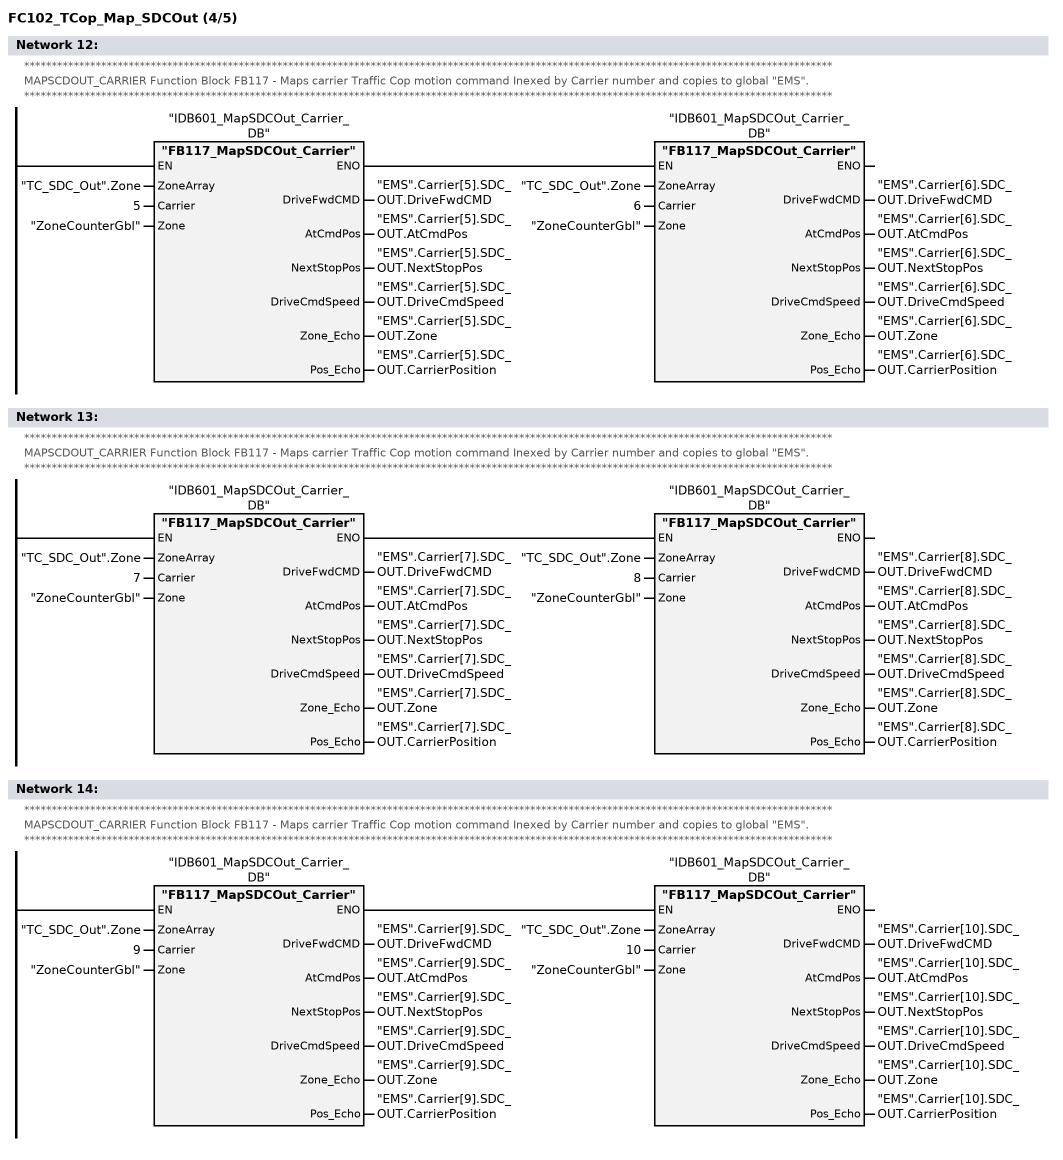
   RUNG wire#powerrail
      "IDB601_MapSDCOut_Carrier_DB"(ZoneArray := "TC_SDC_Out".Zone, Carrier := 5, Zone := "ZoneCounterGbl", DriveFwdCMD => "EMS".Carrier[5].SDC_OUT.DriveFwdCMD, AtCmdPos => "EMS".Carrier[5].SDC_OUT.AtCmdPos, NextStopPos => "EMS".Carrier[5].SDC_OUT.NextStopPos, DriveCmdSpeed => "EMS".Carrier[5].SDC_OUT.DriveCmdSpeed, Zone_Echo => "EMS".Carrier[5].SDC_OUT.Zone, Pos_Echo => "EMS".Carrier[5].SDC_OUT.CarrierPosition)
      "IDB601_MapSDCOut_Carrier_DB"(ZoneArray := "TC_SDC_Out".Zone, Carrier := 6, Zone := "ZoneCounterGbl", DriveFwdCMD => "EMS".Carrier[6].SDC_OUT.DriveFwdCMD, AtCmdPos => "EMS".Carrier[6].SDC_OUT.AtCmdPos, NextStopPos => "EMS".Carrier[6].SDC_OUT.NextStopPos, DriveCmdSpeed => "EMS".Carrier[6].SDC_OUT.DriveCmdSpeed, Zone_Echo => "EMS".Carrier[6].SDC_OUT.Zone, Pos_Echo => "EMS".Carrier[6].SDC_OUT.CarrierPosition)
   END_RUNG
   // the same network as SCL:
   "IDB601_MapSDCOut_Carrier_DB"(ZoneArray := "TC_SDC_Out".Zone,   // "FB117_MapSDCOut_Carrier"
                           Carrier := 5,
                           Zone := "ZoneCounterGbl",
                           DriveFwdCMD => "EMS".Carrier[5].SDC_OUT.DriveFwdCMD,
                           AtCmdPos => "EMS".Carrier[5].SDC_OUT.AtCmdPos,
                           NextStopPos => "EMS".Carrier[5].SDC_OUT.NextStopPos,
                           DriveCmdSpeed => "EMS".Carrier[5].SDC_OUT.DriveCmdSpeed,
                           Zone_Echo => "EMS".Carrier[5].SDC_OUT.Zone,
                           Pos_Echo => "EMS".Carrier[5].SDC_OUT.CarrierPosition,
                           ENO => #_w1);
   IF #_w1 THEN
       "IDB601_MapSDCOut_Carrier_DB"(ZoneArray := "TC_SDC_Out".Zone,   // "FB117_MapSDCOut_Carrier"
                               Carrier := 6,
                               Zone := "ZoneCounterGbl",
                               DriveFwdCMD => "EMS".Carrier[6].SDC_OUT.DriveFwdCMD,
                               AtCmdPos => "EMS".Carrier[6].SDC_OUT.AtCmdPos,
                               NextStopPos => "EMS".Carrier[6].SDC_OUT.NextStopPos,
                               DriveCmdSpeed => "EMS".Carrier[6].SDC_OUT.DriveCmdSpeed,
                               Zone_Echo => "EMS".Carrier[6].SDC_OUT.Zone,
                               Pos_Echo => "EMS".Carrier[6].SDC_OUT.CarrierPosition);
   END_IF;
END_REGION

REGION Network 13
   // ***************************************************************************************************************************************************
   // 
   // MAPSCDOUT_CARRIER Function Block FB117 - Maps carrier Traffic Cop motion command Inexed by Carrier number and copies to global "EMS". 
   // 
   // ***************************************************************************************************************************************************
   RUNG wire#powerrail
      "IDB601_MapSDCOut_Carrier_DB"(ZoneArray := "TC_SDC_Out".Zone, Carrier := 7, Zone := "ZoneCounterGbl", DriveFwdCMD => "EMS".Carrier[7].SDC_OUT.DriveFwdCMD, AtCmdPos => "EMS".Carrier[7].SDC_OUT.AtCmdPos, NextStopPos => "EMS".Carrier[7].SDC_OUT.NextStopPos, DriveCmdSpeed => "EMS".Carrier[7].SDC_OUT.DriveCmdSpeed, Zone_Echo => "EMS".Carrier[7].SDC_OUT.Zone, Pos_Echo => "EMS".Carrier[7].SDC_OUT.CarrierPosition)
      "IDB601_MapSDCOut_Carrier_DB"(ZoneArray := "TC_SDC_Out".Zone, Carrier := 8, Zone := "ZoneCounterGbl", DriveFwdCMD => "EMS".Carrier[8].SDC_OUT.DriveFwdCMD, AtCmdPos => "EMS".Carrier[8].SDC_OUT.AtCmdPos, NextStopPos => "EMS".Carrier[8].SDC_OUT.NextStopPos, DriveCmdSpeed => "EMS".Carrier[8].SDC_OUT.DriveCmdSpeed, Zone_Echo => "EMS".Carrier[8].SDC_OUT.Zone, Pos_Echo => "EMS".Carrier[8].SDC_OUT.CarrierPosition)
   END_RUNG
   // the same network as SCL:
   "IDB601_MapSDCOut_Carrier_DB"(ZoneArray := "TC_SDC_Out".Zone,   // "FB117_MapSDCOut_Carrier"
                           Carrier := 7,
                           Zone := "ZoneCounterGbl",
                           DriveFwdCMD => "EMS".Carrier[7].SDC_OUT.DriveFwdCMD,
                           AtCmdPos => "EMS".Carrier[7].SDC_OUT.AtCmdPos,
                           NextStopPos => "EMS".Carrier[7].SDC_OUT.NextStopPos,
                           DriveCmdSpeed => "EMS".Carrier[7].SDC_OUT.DriveCmdSpeed,
                           Zone_Echo => "EMS".Carrier[7].SDC_OUT.Zone,
                           Pos_Echo => "EMS".Carrier[7].SDC_OUT.CarrierPosition,
                           ENO => #_w1);
   IF #_w1 THEN
       "IDB601_MapSDCOut_Carrier_DB"(ZoneArray := "TC_SDC_Out".Zone,   // "FB117_MapSDCOut_Carrier"
                               Carrier := 8,
                               Zone := "ZoneCounterGbl",
                               DriveFwdCMD => "EMS".Carrier[8].SDC_OUT.DriveFwdCMD,
                               AtCmdPos => "EMS".Carrier[8].SDC_OUT.AtCmdPos,
                               NextStopPos => "EMS".Carrier[8].SDC_OUT.NextStopPos,
                               DriveCmdSpeed => "EMS".Carrier[8].SDC_OUT.DriveCmdSpeed,
                               Zone_Echo => "EMS".Carrier[8].SDC_OUT.Zone,
                               Pos_Echo => "EMS".Carrier[8].SDC_OUT.CarrierPosition);
   END_IF;
END_REGION

REGION Network 14
   // ***************************************************************************************************************************************************
   // 
   // MAPSCDOUT_CARRIER Function Block FB117 - Maps carrier Traffic Cop motion command Inexed by Carrier number and copies to global "EMS". 
   // 
   // ***************************************************************************************************************************************************
   RUNG wire#powerrail
      "IDB601_MapSDCOut_Carrier_DB"(ZoneArray := "TC_SDC_Out".Zone, Carrier := 9, Zone := "ZoneCounterGbl", DriveFwdCMD => "EMS".Carrier[9].SDC_OUT.DriveFwdCMD, AtCmdPos => "EMS".Carrier[9].SDC_OUT.AtCmdPos, NextStopPos => "EMS".Carrier[9].SDC_OUT.NextStopPos, DriveCmdSpeed => "EMS".Carrier[9].SDC_OUT.DriveCmdSpeed, Zone_Echo => "EMS".Carrier[9].SDC_OUT.Zone, Pos_Echo => "EMS".Carrier[9].SDC_OUT.CarrierPosition)
      "IDB601_MapSDCOut_Carrier_DB"(ZoneArray := "TC_SDC_Out".Zone, Carrier := 10, Zone := "ZoneCounterGbl", DriveFwdCMD => "EMS".Carrier[10].SDC_OUT.DriveFwdCMD, AtCmdPos => "EMS".Carrier[10].SDC_OUT.AtCmdPos, NextStopPos => "EMS".Carrier[10].SDC_OUT.NextStopPos, DriveCmdSpeed => "EMS".Carrier[10].SDC_OUT.DriveCmdSpeed, Zone_Echo => "EMS".Carrier[10].SDC_OUT.Zone, Pos_Echo => "EMS".Carrier[10].SDC_OUT.CarrierPosition)
   END_RUNG
   // the same network as SCL:
   "IDB601_MapSDCOut_Carrier_DB"(ZoneArray := "TC_SDC_Out".Zone,   // "FB117_MapSDCOut_Carrier"
                           Carrier := 9,
                           Zone := "ZoneCounterGbl",
                           DriveFwdCMD => "EMS".Carrier[9].SDC_OUT.DriveFwdCMD,
                           AtCmdPos => "EMS".Carrier[9].SDC_OUT.AtCmdPos,
                           NextStopPos => "EMS".Carrier[9].SDC_OUT.NextStopPos,
                           DriveCmdSpeed => "EMS".Carrier[9].SDC_OUT.DriveCmdSpeed,
                           Zone_Echo => "EMS".Carrier[9].SDC_OUT.Zone,
                           Pos_Echo => "EMS".Carrier[9].SDC_OUT.CarrierPosition,
                           ENO => #_w1);
   IF #_w1 THEN
       "IDB601_MapSDCOut_Carrier_DB"(ZoneArray := "TC_SDC_Out".Zone,   // "FB117_MapSDCOut_Carrier"
                               Carrier := 10,
                               Zone := "ZoneCounterGbl",
                               DriveFwdCMD => "EMS".Carrier[10].SDC_OUT.DriveFwdCMD,
                               AtCmdPos => "EMS".Carrier[10].SDC_OUT.AtCmdPos,
                               NextStopPos => "EMS".Carrier[10].SDC_OUT.NextStopPos,
                               DriveCmdSpeed => "EMS".Carrier[10].SDC_OUT.DriveCmdSpeed,
                               Zone_Echo => "EMS".Carrier[10].SDC_OUT.Zone,
                               Pos_Echo => "EMS".Carrier[10].SDC_OUT.CarrierPosition);
   END_IF;
END_REGION

REGION Network 15
   // ***************************************************************************************************************************************************
   // 
   // MAPSCDOUT_CARRIER Function Block FB117 - Maps carrier Traffic Cop motion command Inexed by Carrier number and copies to global "EMS". 
   // 
   // ***************************************************************************************************************************************************
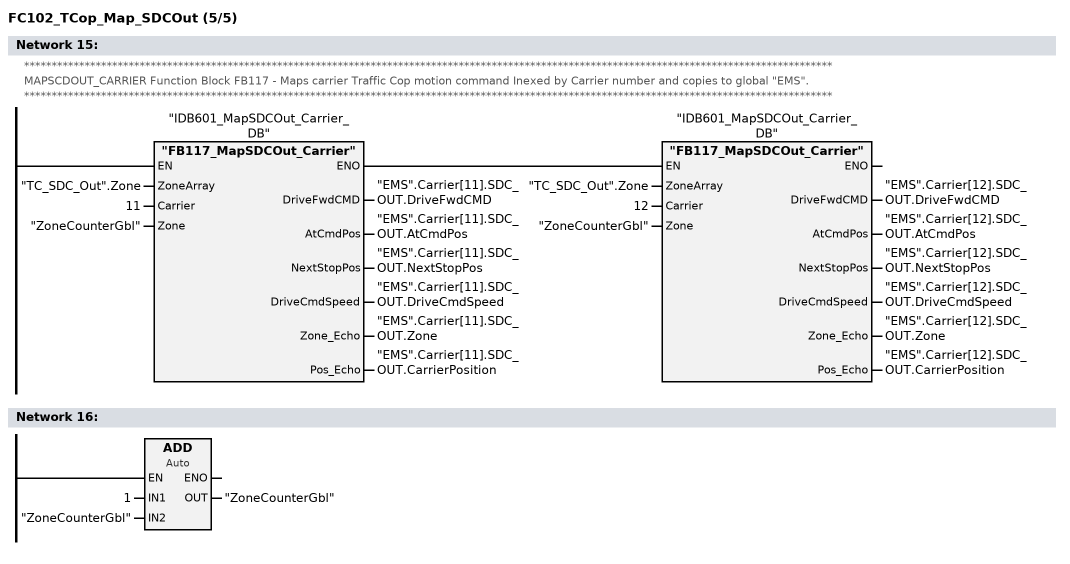
   RUNG wire#powerrail
      "IDB601_MapSDCOut_Carrier_DB"(ZoneArray := "TC_SDC_Out".Zone, Carrier := 11, Zone := "ZoneCounterGbl", DriveFwdCMD => "EMS".Carrier[11].SDC_OUT.DriveFwdCMD, AtCmdPos => "EMS".Carrier[11].SDC_OUT.AtCmdPos, NextStopPos => "EMS".Carrier[11].SDC_OUT.NextStopPos, DriveCmdSpeed => "EMS".Carrier[11].SDC_OUT.DriveCmdSpeed, Zone_Echo => "EMS".Carrier[11].SDC_OUT.Zone, Pos_Echo => "EMS".Carrier[11].SDC_OUT.CarrierPosition)
      "IDB601_MapSDCOut_Carrier_DB"(ZoneArray := "TC_SDC_Out".Zone, Carrier := 12, Zone := "ZoneCounterGbl", DriveFwdCMD => "EMS".Carrier[12].SDC_OUT.DriveFwdCMD, AtCmdPos => "EMS".Carrier[12].SDC_OUT.AtCmdPos, NextStopPos => "EMS".Carrier[12].SDC_OUT.NextStopPos, DriveCmdSpeed => "EMS".Carrier[12].SDC_OUT.DriveCmdSpeed, Zone_Echo => "EMS".Carrier[12].SDC_OUT.Zone, Pos_Echo => "EMS".Carrier[12].SDC_OUT.CarrierPosition)
   END_RUNG
   // the same network as SCL:
   "IDB601_MapSDCOut_Carrier_DB"(ZoneArray := "TC_SDC_Out".Zone,   // "FB117_MapSDCOut_Carrier"
                           Carrier := 11,
                           Zone := "ZoneCounterGbl",
                           DriveFwdCMD => "EMS".Carrier[11].SDC_OUT.DriveFwdCMD,
                           AtCmdPos => "EMS".Carrier[11].SDC_OUT.AtCmdPos,
                           NextStopPos => "EMS".Carrier[11].SDC_OUT.NextStopPos,
                           DriveCmdSpeed => "EMS".Carrier[11].SDC_OUT.DriveCmdSpeed,
                           Zone_Echo => "EMS".Carrier[11].SDC_OUT.Zone,
                           Pos_Echo => "EMS".Carrier[11].SDC_OUT.CarrierPosition,
                           ENO => #_w1);
   IF #_w1 THEN
       "IDB601_MapSDCOut_Carrier_DB"(ZoneArray := "TC_SDC_Out".Zone,   // "FB117_MapSDCOut_Carrier"
                               Carrier := 12,
                               Zone := "ZoneCounterGbl",
                               DriveFwdCMD => "EMS".Carrier[12].SDC_OUT.DriveFwdCMD,
                               AtCmdPos => "EMS".Carrier[12].SDC_OUT.AtCmdPos,
                               NextStopPos => "EMS".Carrier[12].SDC_OUT.NextStopPos,
                               DriveCmdSpeed => "EMS".Carrier[12].SDC_OUT.DriveCmdSpeed,
                               Zone_Echo => "EMS".Carrier[12].SDC_OUT.Zone,
                               Pos_Echo => "EMS".Carrier[12].SDC_OUT.CarrierPosition);
   END_IF;
END_REGION

REGION Network 16
   RUNG wire#powerrail
      Add(in1 := 1, in2 := "ZoneCounterGbl", out => "ZoneCounterGbl")
   END_RUNG
   // the same network as SCL:
   "ZoneCounterGbl" := 1 + "ZoneCounterGbl";
END_REGION
END_FUNCTION

FUNCTION "FC103_SystemZoneFind" : Void   // FC103, LAD
{ S7_Optimized_Access := 'FALSE' }
VERSION : 0.1
   VAR_TEMP
      resettemp : Bool;
      dntemp : Bool;
   END_VAR
BEGIN

REGION Network 1
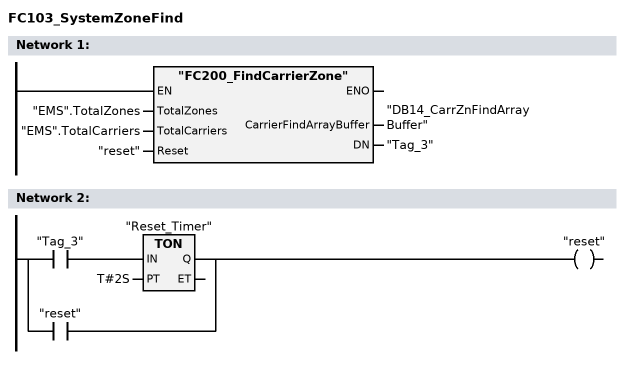
   RUNG wire#powerrail
      "FC200_FindCarrierZone"(TotalZones := "EMS".TotalZones, TotalCarriers := "EMS".TotalCarriers, Reset := "reset", CarrierFindArrayBuffer => "DB14_CarrZnFindArrayBuffer", DN => "Tag_3")
   END_RUNG
   // the same network as SCL:
   "FC200_FindCarrierZone"(TotalZones := "EMS".TotalZones,
                           TotalCarriers := "EMS".TotalCarriers,
                           Reset := "reset",
                           CarrierFindArrayBuffer => "DB14_CarrZnFindArrayBuffer",
                           DN => "Tag_3");
END_REGION

REGION Network 2
   "Reset_Timer".TON(IN := "Tag_3", PT := T#2S);
   "reset" := "Reset_Timer".Q OR "reset";
END_REGION
END_FUNCTION

FUNCTION "FC104_CarrierSetup" : Void   // FC104, LAD
{ S7_Optimized_Access := 'FALSE' }
VERSION : 0.1
   VAR_TEMP
      CarrierCounter : Int;
      TotalCarriers : Int;
      CounterReset : Bool;
      CarrierCounterDN : Bool;
      OneShotClock_2hz : Bool;
   END_VAR
BEGIN

REGION Network 1
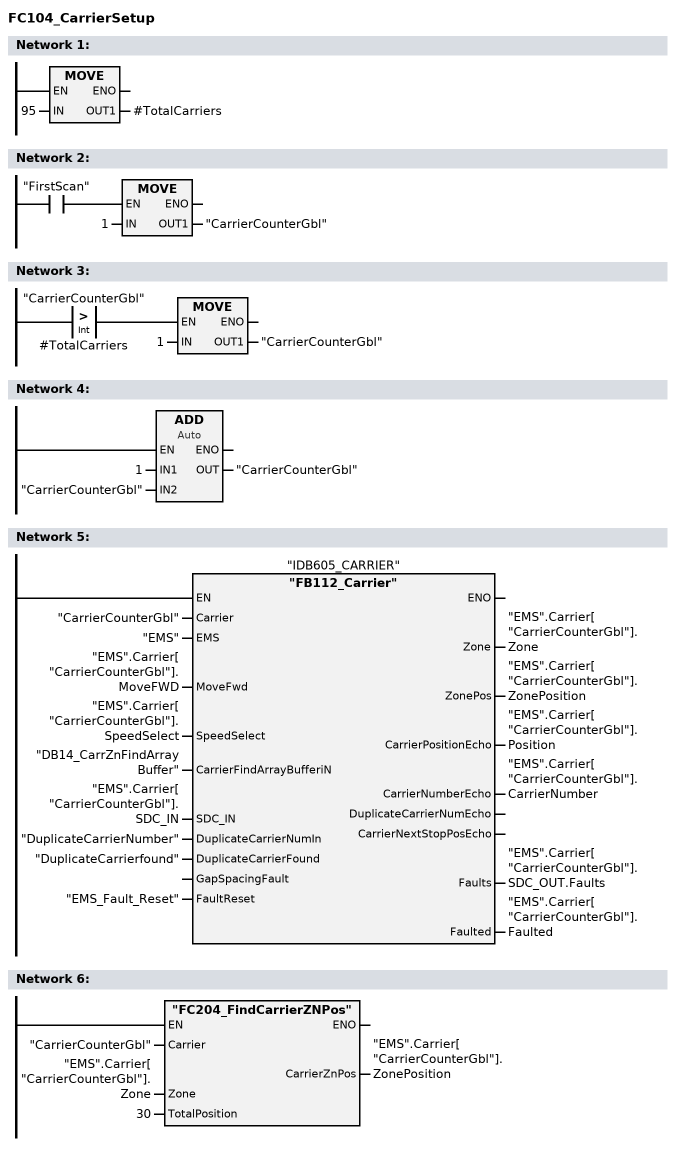
   RUNG wire#powerrail
      Move(in := 95, out1 => #TotalCarriers)
   END_RUNG
   // the same network as SCL:
   #TotalCarriers := 95;
END_REGION

REGION Network 2
   RUNG wire#powerrail
      Contact( "FirstScan" )
      Move(in := 1, out1 => "CarrierCounterGbl")
   END_RUNG
   // the same network as SCL:
   IF "FirstScan" THEN "CarrierCounterGbl" := 1; END_IF;
END_REGION

REGION Network 3
   RUNG wire#powerrail
      { S7_Templates := "SrcType := Int" } GT_Contact(in1 := "CarrierCounterGbl", in2 := #TotalCarriers)
      Move(in := 1, out1 => "CarrierCounterGbl")
   END_RUNG
   // the same network as SCL:
   IF "CarrierCounterGbl" > #TotalCarriers THEN "CarrierCounterGbl" := 1; END_IF;
END_REGION

REGION Network 4
   RUNG wire#powerrail
      Add(in1 := 1, in2 := "CarrierCounterGbl", out => "CarrierCounterGbl")
   END_RUNG
   // the same network as SCL:
   "CarrierCounterGbl" := 1 + "CarrierCounterGbl";
END_REGION

REGION Network 5
   RUNG wire#powerrail
      "IDB605_CARRIER"(Carrier := "CarrierCounterGbl", EMS := "EMS", MoveFwd := "EMS".Carrier["CarrierCounterGbl"].MoveFWD, SpeedSelect := "EMS".Carrier["CarrierCounterGbl"].SpeedSelect, CarrierFindArrayBufferiN := "DB14_CarrZnFindArrayBuffer", SDC_IN := "EMS".Carrier["CarrierCounterGbl"].SDC_IN, DuplicateCarrierNumIn := "DuplicateCarrierNumber", DuplicateCarrierFound := "DuplicateCarrierfound", GapSpacingFault :=, FaultReset := "EMS_Fault_Reset", Zone => "EMS".Carrier["CarrierCounterGbl"].Zone, ZonePos => "EMS".Carrier["CarrierCounterGbl"].ZonePosition, CarrierPositionEcho => "EMS".Carrier["CarrierCounterGbl"].Position, CarrierNumberEcho => "EMS".Carrier["CarrierCounterGbl"].CarrierNumber, DuplicateCarrierNumEcho =>, CarrierNextStopPosEcho =>, Faults => "EMS".Carrier["CarrierCounterGbl"].SDC_OUT.Faults, Faulted => "EMS".Carrier["CarrierCounterGbl"].Faulted)
   END_RUNG
   // the same network as SCL:
   "IDB605_CARRIER"(Carrier := "CarrierCounterGbl",   // "FB112_Carrier"
                    EMS := "EMS",
                    MoveFwd := "EMS".Carrier["CarrierCounterGbl"].MoveFWD,
                    SpeedSelect := "EMS".Carrier["CarrierCounterGbl"].SpeedSelect,
                    CarrierFindArrayBufferiN := "DB14_CarrZnFindArrayBuffer",
                    SDC_IN := "EMS".Carrier["CarrierCounterGbl"].SDC_IN,
                    DuplicateCarrierNumIn := "DuplicateCarrierNumber",
                    DuplicateCarrierFound := "DuplicateCarrierfound",
                    FaultReset := "EMS_Fault_Reset",
                    Zone => "EMS".Carrier["CarrierCounterGbl"].Zone,
                    ZonePos => "EMS".Carrier["CarrierCounterGbl"].ZonePosition,
                    CarrierPositionEcho => "EMS".Carrier["CarrierCounterGbl"].Position,
                    CarrierNumberEcho => "EMS".Carrier["CarrierCounterGbl"].CarrierNumber,
                    Faults => "EMS".Carrier["CarrierCounterGbl"].SDC_OUT.Faults,
                    Faulted => "EMS".Carrier["CarrierCounterGbl"].Faulted);
END_REGION

REGION Network 6
   RUNG wire#powerrail
      "FC204_FindCarrierZNPos"(Carrier := "CarrierCounterGbl", Zone := "EMS".Carrier["CarrierCounterGbl"].Zone, TotalPosition := 30, CarrierZnPos => "EMS".Carrier["CarrierCounterGbl"].ZonePosition)
   END_RUNG
   // the same network as SCL:
   "FC204_FindCarrierZNPos"(Carrier := "CarrierCounterGbl",
                           Zone := "EMS".Carrier["CarrierCounterGbl"].Zone,
                           TotalPosition := 30,
                           CarrierZnPos => "EMS".Carrier["CarrierCounterGbl"].ZonePosition);
END_REGION
END_FUNCTION

FUNCTION "FC105_EMS_State" : Void   // FC105, SCL
{ S7_Optimized_Access := 'TRUE' }
VERSION : 0.1
   VAR_TEMP
      N : Int;
   END_VAR
BEGIN
   FOR #N := 1 TO 82 DO
       // Statement section FOR
       IF "DB16_EMS_Status".EMS_DeviceStates.DeviceStates_State4[#N] = FALSE
       THEN
           "DB16_EMS_Status".EMS_DeviceStates.DeviceStates_Condition_HMI[#N] := 0;
       ELSE
           IF "DB16_EMS_Status".EMS_DeviceStates.DeviceStates_State4[#N] = TRUE
           THEN
               "DB16_EMS_Status".EMS_DeviceStates.DeviceStates_Condition_HMI[#N] := 1;
           END_IF;
           IF "DB16_EMS_Status".EMS_DeviceStates.DeviceStates_State5[#N] = TRUE
           THEN
               "DB16_EMS_Status".EMS_DeviceStates.DeviceStates_Condition_HMI[#N] := 3;
           END_IF;
           IF "DB16_EMS_Status".EMS_DeviceStates.DeviceStates_State2[#N] = TRUE
           THEN
               "DB16_EMS_Status".EMS_DeviceStates.DeviceStates_Condition_HMI[#N] := 2;
           END_IF;
       END_IF;

   END_FOR;
END_FUNCTION

FUNCTION "FC106_SDC_To_Carrier_Map_IO [C01-C10]" : Void   // FC106, LAD
{ S7_Optimized_Access := 'TRUE' }
VERSION : 0.1
   VAR_TEMP
      templatch : Bool;
   END_VAR
BEGIN

REGION Network 1
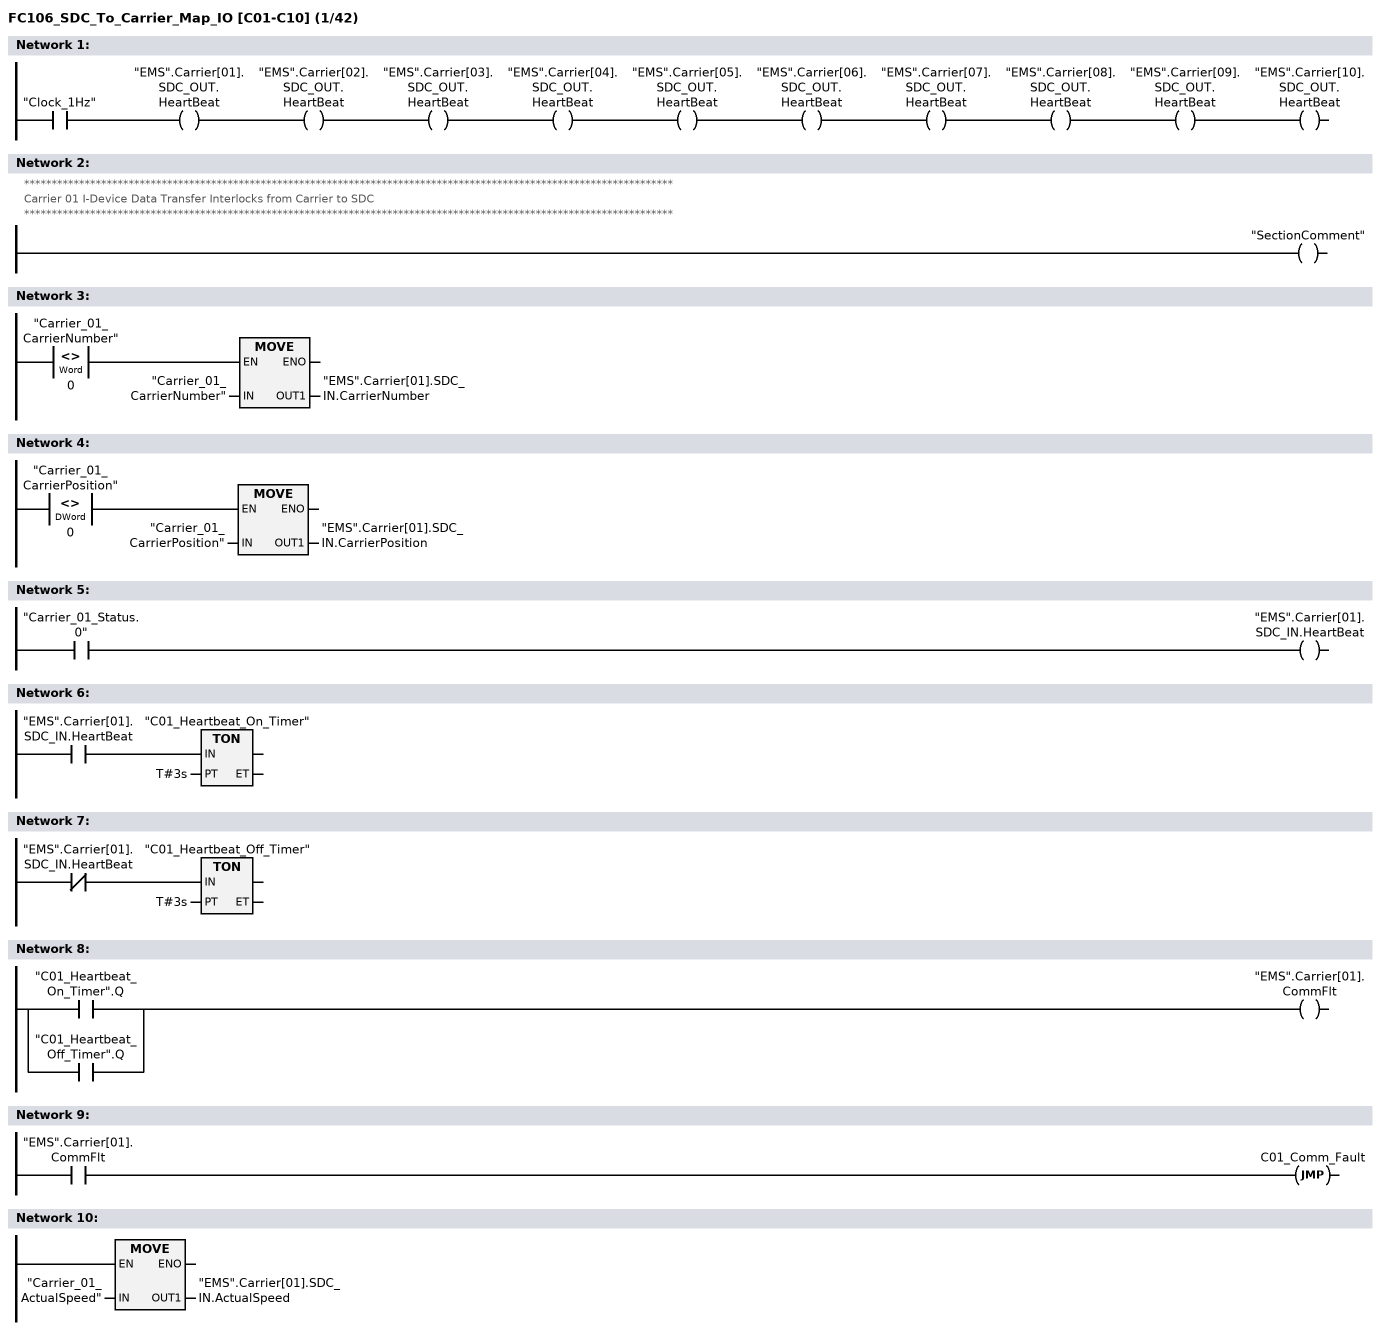
   RUNG wire#powerrail
      Contact( "Clock_1Hz" )
      Coil( "EMS".Carrier[01].SDC_OUT.HeartBeat )
      Coil( "EMS".Carrier[02].SDC_OUT.HeartBeat )
      Coil( "EMS".Carrier[03].SDC_OUT.HeartBeat )
      Coil( "EMS".Carrier[04].SDC_OUT.HeartBeat )
      Coil( "EMS".Carrier[05].SDC_OUT.HeartBeat )
      Coil( "EMS".Carrier[06].SDC_OUT.HeartBeat )
      Coil( "EMS".Carrier[07].SDC_OUT.HeartBeat )
      Coil( "EMS".Carrier[08].SDC_OUT.HeartBeat )
      Coil( "EMS".Carrier[09].SDC_OUT.HeartBeat )
      Coil( "EMS".Carrier[10].SDC_OUT.HeartBeat )
   END_RUNG
   // the same network as SCL:
   "EMS".Carrier[01].SDC_OUT.HeartBeat := "Clock_1Hz";
   "EMS".Carrier[02].SDC_OUT.HeartBeat := "Clock_1Hz";
   "EMS".Carrier[03].SDC_OUT.HeartBeat := "Clock_1Hz";
   "EMS".Carrier[04].SDC_OUT.HeartBeat := "Clock_1Hz";
   "EMS".Carrier[05].SDC_OUT.HeartBeat := "Clock_1Hz";
   "EMS".Carrier[06].SDC_OUT.HeartBeat := "Clock_1Hz";
   "EMS".Carrier[07].SDC_OUT.HeartBeat := "Clock_1Hz";
   "EMS".Carrier[08].SDC_OUT.HeartBeat := "Clock_1Hz";
   "EMS".Carrier[09].SDC_OUT.HeartBeat := "Clock_1Hz";
   "EMS".Carrier[10].SDC_OUT.HeartBeat := "Clock_1Hz";
END_REGION

REGION Network 2
   // **********************************************************************************************************************
   // 
   // Carrier 01 I-Device Data Transfer Interlocks from Carrier to SDC
   // 
   // **********************************************************************************************************************
   RUNG wire#powerrail
      Coil( "SectionComment" )
   END_RUNG
   // the same network as SCL:
   "SectionComment" := TRUE;
END_REGION

REGION Network 3
   RUNG wire#powerrail
      { S7_Templates := "SrcType := Word" } NE_Contact(in1 := "Carrier_01_CarrierNumber", in2 := 0)
      Move(in := "Carrier_01_CarrierNumber", out1 => "EMS".Carrier[01].SDC_IN.CarrierNumber)
   END_RUNG
   // the same network as SCL:
   IF "Carrier_01_CarrierNumber" <> 0 THEN
       "EMS".Carrier[01].SDC_IN.CarrierNumber := "Carrier_01_CarrierNumber";
   END_IF;
END_REGION

REGION Network 4
   RUNG wire#powerrail
      { S7_Templates := "SrcType := DWord" } NE_Contact(in1 := "Carrier_01_CarrierPosition", in2 := 0)
      Move(in := "Carrier_01_CarrierPosition", out1 => "EMS".Carrier[01].SDC_IN.CarrierPosition)
   END_RUNG
   // the same network as SCL:
   IF "Carrier_01_CarrierPosition" <> 0 THEN
       "EMS".Carrier[01].SDC_IN.CarrierPosition := "Carrier_01_CarrierPosition";
   END_IF;
END_REGION

REGION Network 5
   RUNG wire#powerrail
      Contact( "Carrier_01_Status.0" )
      Coil( "EMS".Carrier[01].SDC_IN.HeartBeat )
   END_RUNG
   // the same network as SCL:
   "EMS".Carrier[01].SDC_IN.HeartBeat := "Carrier_01_Status.0";
END_REGION

REGION Network 6
   "C01_Heartbeat_On_Timer".TON(IN := "EMS".Carrier[01].SDC_IN.HeartBeat, PT := T#3s);
END_REGION

REGION Network 7
   "C01_Heartbeat_Off_Timer".TON(IN := NOT "EMS".Carrier[01].SDC_IN.HeartBeat, PT := T#3s);
END_REGION

REGION Network 8
   RUNG wire#powerrail
      Contact( "C01_Heartbeat_On_Timer".Q )
      wire#w1
      Coil( "EMS".Carrier[01].CommFlt )
   END_RUNG
   RUNG wire#powerrail
      Contact( "C01_Heartbeat_Off_Timer".Q )
   END_RUNG wire#w1
   // the same network as SCL:
   "EMS".Carrier[01].CommFlt := "C01_Heartbeat_On_Timer".Q OR "C01_Heartbeat_Off_Timer".Q;
END_REGION

REGION Network 9
   RUNG wire#powerrail
      Contact( "EMS".Carrier[01].CommFlt )
      JumpCoil( C01_Comm_Fault )
   END_RUNG
   // the same network as SCL:
   IF "EMS".Carrier[01].CommFlt THEN GOTO C01_Comm_Fault; END_IF;
END_REGION

REGION Network 10
   RUNG wire#powerrail
      Move(in := "Carrier_01_ActualSpeed", out1 => "EMS".Carrier[01].SDC_IN.ActualSpeed)
   END_RUNG
   // the same network as SCL:
   "EMS".Carrier[01].SDC_IN.ActualSpeed := "Carrier_01_ActualSpeed";
END_REGION

REGION Network 11
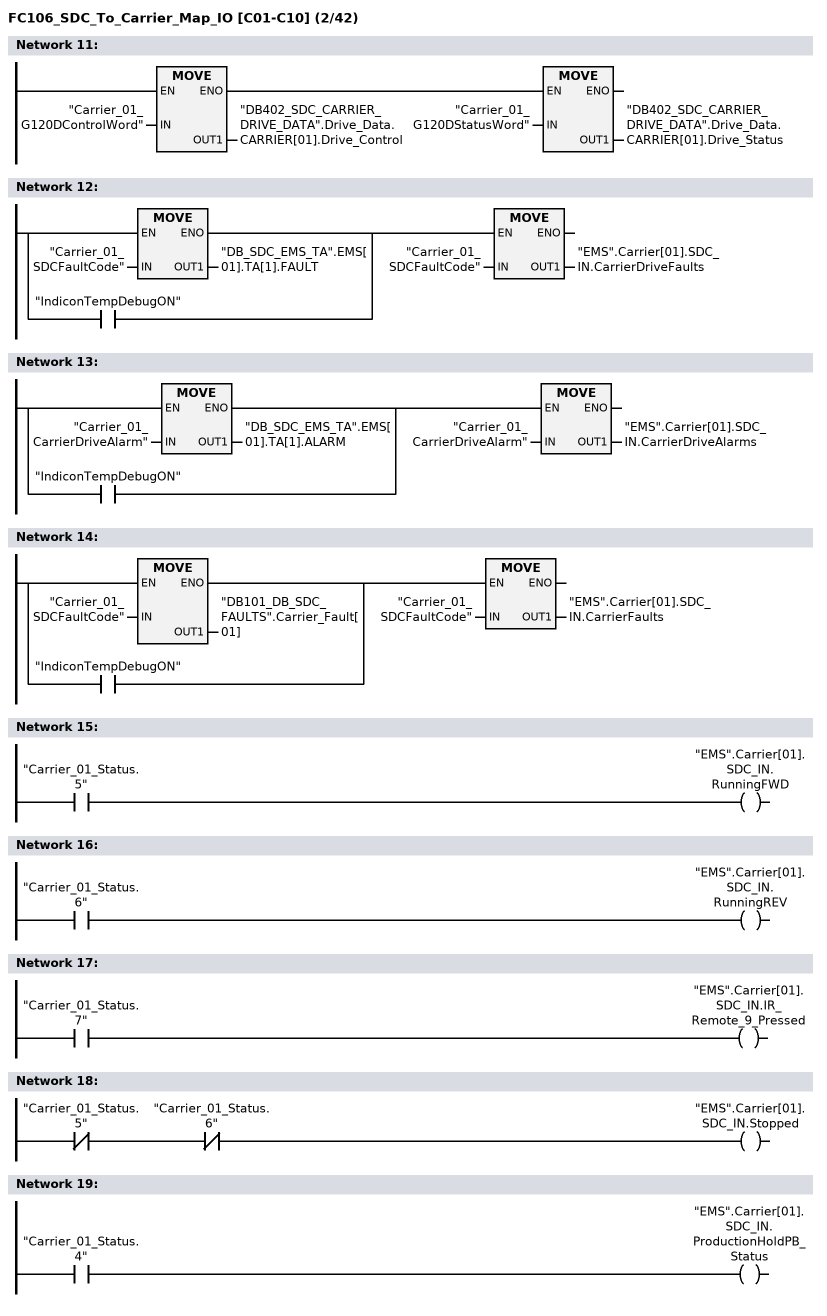
   RUNG wire#powerrail
      Move(in := "Carrier_01_G120DControlWord", out1 => "DB402_SDC_CARRIER_DRIVE_DATA".Drive_Data.CARRIER[01].Drive_Control)
      Move(in := "Carrier_01_G120DStatusWord", out1 => "DB402_SDC_CARRIER_DRIVE_DATA".Drive_Data.CARRIER[01].Drive_Status)
   END_RUNG
   // the same network as SCL:
   "DB402_SDC_CARRIER_DRIVE_DATA".Drive_Data.CARRIER[01].Drive_Control := "Carrier_01_G120DControlWord";
   "DB402_SDC_CARRIER_DRIVE_DATA".Drive_Data.CARRIER[01].Drive_Status := "Carrier_01_G120DStatusWord";
END_REGION

REGION Network 12
   RUNG wire#powerrail
      Move(in := "Carrier_01_SDCFaultCode", out1 => "DB_SDC_EMS_TA".EMS[01].TA[1].FAULT)
      wire#w1
      Move(in := "Carrier_01_SDCFaultCode", out1 => "EMS".Carrier[01].SDC_IN.CarrierDriveFaults)
   END_RUNG
   RUNG wire#powerrail
      Contact( "IndiconTempDebugON" )
   END_RUNG wire#w1
   // the same network as SCL:
   "DB_SDC_EMS_TA".EMS[01].TA[1].FAULT := "Carrier_01_SDCFaultCode";
   IF TRUE OR "IndiconTempDebugON" THEN
       "EMS".Carrier[01].SDC_IN.CarrierDriveFaults := "Carrier_01_SDCFaultCode";
   END_IF;
END_REGION

REGION Network 13
   RUNG wire#powerrail
      Move(in := "Carrier_01_CarrierDriveAlarm", out1 => "DB_SDC_EMS_TA".EMS[01].TA[1].ALARM)
      wire#w1
      Move(in := "Carrier_01_CarrierDriveAlarm", out1 => "EMS".Carrier[01].SDC_IN.CarrierDriveAlarms)
   END_RUNG
   RUNG wire#powerrail
      Contact( "IndiconTempDebugON" )
   END_RUNG wire#w1
   // the same network as SCL:
   "DB_SDC_EMS_TA".EMS[01].TA[1].ALARM := "Carrier_01_CarrierDriveAlarm";
   IF TRUE OR "IndiconTempDebugON" THEN
       "EMS".Carrier[01].SDC_IN.CarrierDriveAlarms := "Carrier_01_CarrierDriveAlarm";
   END_IF;
END_REGION

REGION Network 14
   RUNG wire#powerrail
      Move(in := "Carrier_01_SDCFaultCode", out1 => "DB101_DB_SDC_FAULTS".Carrier_Fault[01])
      wire#w1
      Move(in := "Carrier_01_SDCFaultCode", out1 => "EMS".Carrier[01].SDC_IN.CarrierFaults)
   END_RUNG
   RUNG wire#powerrail
      Contact( "IndiconTempDebugON" )
   END_RUNG wire#w1
   // the same network as SCL:
   "DB101_DB_SDC_FAULTS".Carrier_Fault[01] := "Carrier_01_SDCFaultCode";
   IF TRUE OR "IndiconTempDebugON" THEN
       "EMS".Carrier[01].SDC_IN.CarrierFaults := "Carrier_01_SDCFaultCode";
   END_IF;
END_REGION

REGION Network 15
   RUNG wire#powerrail
      Contact( "Carrier_01_Status.5" )
      Coil( "EMS".Carrier[01].SDC_IN.RunningFWD )
   END_RUNG
   // the same network as SCL:
   "EMS".Carrier[01].SDC_IN.RunningFWD := "Carrier_01_Status.5";
END_REGION

REGION Network 16
   RUNG wire#powerrail
      Contact( "Carrier_01_Status.6" )
      Coil( "EMS".Carrier[01].SDC_IN.RunningREV )
   END_RUNG
   // the same network as SCL:
   "EMS".Carrier[01].SDC_IN.RunningREV := "Carrier_01_Status.6";
END_REGION

REGION Network 17
   RUNG wire#powerrail
      Contact( "Carrier_01_Status.7" )
      Coil( "EMS".Carrier[01].SDC_IN.IR_Remote_9_Pressed )
   END_RUNG
   // the same network as SCL:
   "EMS".Carrier[01].SDC_IN.IR_Remote_9_Pressed := "Carrier_01_Status.7";
END_REGION

REGION Network 18
   RUNG wire#powerrail
      I_Contact( "Carrier_01_Status.5" )
      I_Contact( "Carrier_01_Status.6" )
      Coil( "EMS".Carrier[01].SDC_IN.Stopped )
   END_RUNG
   // the same network as SCL:
   "EMS".Carrier[01].SDC_IN.Stopped := NOT "Carrier_01_Status.5" AND NOT "Carrier_01_Status.6";
END_REGION

REGION Network 19
   RUNG wire#powerrail
      Contact( "Carrier_01_Status.4" )
      Coil( "EMS".Carrier[01].SDC_IN.ProductionHoldPB_Status )
   END_RUNG
   // the same network as SCL:
   "EMS".Carrier[01].SDC_IN.ProductionHoldPB_Status := "Carrier_01_Status.4";
END_REGION

REGION Network 20
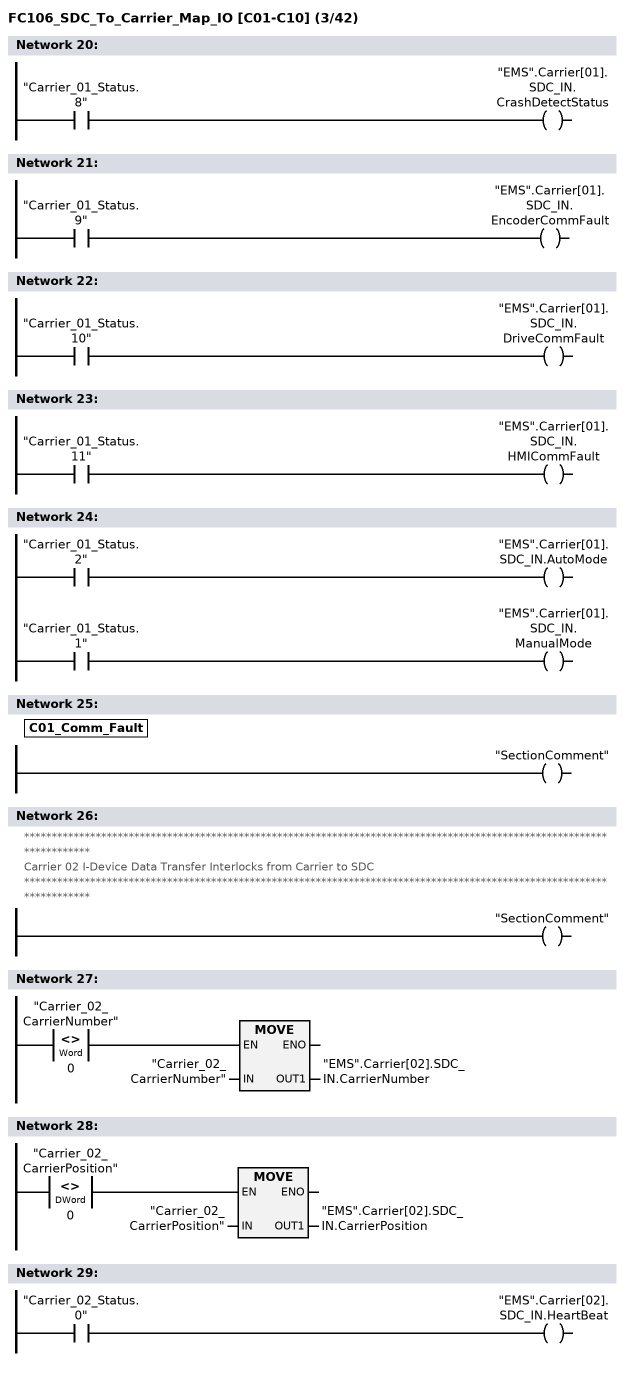
   RUNG wire#powerrail
      Contact( "Carrier_01_Status.8" )
      Coil( "EMS".Carrier[01].SDC_IN.CrashDetectStatus )
   END_RUNG
   // the same network as SCL:
   "EMS".Carrier[01].SDC_IN.CrashDetectStatus := "Carrier_01_Status.8";
END_REGION

REGION Network 21
   RUNG wire#powerrail
      Contact( "Carrier_01_Status.9" )
      Coil( "EMS".Carrier[01].SDC_IN.EncoderCommFault )
   END_RUNG
   // the same network as SCL:
   "EMS".Carrier[01].SDC_IN.EncoderCommFault := "Carrier_01_Status.9";
END_REGION

REGION Network 22
   RUNG wire#powerrail
      Contact( "Carrier_01_Status.10" )
      Coil( "EMS".Carrier[01].SDC_IN.DriveCommFault )
   END_RUNG
   // the same network as SCL:
   "EMS".Carrier[01].SDC_IN.DriveCommFault := "Carrier_01_Status.10";
END_REGION

REGION Network 23
   RUNG wire#powerrail
      Contact( "Carrier_01_Status.11" )
      Coil( "EMS".Carrier[01].SDC_IN.HMICommFault )
   END_RUNG
   // the same network as SCL:
   "EMS".Carrier[01].SDC_IN.HMICommFault := "Carrier_01_Status.11";
END_REGION

REGION Network 24
   RUNG wire#powerrail
      Contact( "Carrier_01_Status.2" )
      Coil( "EMS".Carrier[01].SDC_IN.AutoMode )
   END_RUNG
   RUNG wire#powerrail
      Contact( "Carrier_01_Status.1" )
      Coil( "EMS".Carrier[01].SDC_IN.ManualMode )
   END_RUNG
   // the same network as SCL:
   "EMS".Carrier[01].SDC_IN.AutoMode := "Carrier_01_Status.2";
   "EMS".Carrier[01].SDC_IN.ManualMode := "Carrier_01_Status.1";
END_REGION

REGION Network 25
   Label( C01_Comm_Fault )
   RUNG wire#powerrail
      Coil( "SectionComment" )
   END_RUNG
   // the same network as SCL:
   C01_Comm_Fault:
   "SectionComment" := TRUE;
END_REGION

REGION Network 26
   // **********************************************************************************************************************
   // 
   // Carrier 02 I-Device Data Transfer Interlocks from Carrier to SDC
   // 
   // **********************************************************************************************************************
   RUNG wire#powerrail
      Coil( "SectionComment" )
   END_RUNG
   // the same network as SCL:
   "SectionComment" := TRUE;
END_REGION

REGION Network 27
   RUNG wire#powerrail
      { S7_Templates := "SrcType := Word" } NE_Contact(in1 := "Carrier_02_CarrierNumber", in2 := 0)
      Move(in := "Carrier_02_CarrierNumber", out1 => "EMS".Carrier[02].SDC_IN.CarrierNumber)
   END_RUNG
   // the same network as SCL:
   IF "Carrier_02_CarrierNumber" <> 0 THEN
       "EMS".Carrier[02].SDC_IN.CarrierNumber := "Carrier_02_CarrierNumber";
   END_IF;
END_REGION

REGION Network 28
   RUNG wire#powerrail
      { S7_Templates := "SrcType := DWord" } NE_Contact(in1 := "Carrier_02_CarrierPosition", in2 := 0)
      Move(in := "Carrier_02_CarrierPosition", out1 => "EMS".Carrier[02].SDC_IN.CarrierPosition)
   END_RUNG
   // the same network as SCL:
   IF "Carrier_02_CarrierPosition" <> 0 THEN
       "EMS".Carrier[02].SDC_IN.CarrierPosition := "Carrier_02_CarrierPosition";
   END_IF;
END_REGION

REGION Network 29
   RUNG wire#powerrail
      Contact( "Carrier_02_Status.0" )
      Coil( "EMS".Carrier[02].SDC_IN.HeartBeat )
   END_RUNG
   // the same network as SCL:
   "EMS".Carrier[02].SDC_IN.HeartBeat := "Carrier_02_Status.0";
END_REGION

REGION Network 30